(* Logix 5000 project; controller _GigaDiscovery vendor 1 type 14 code 244 rev 35.11; software revision 35.03; part 3 of 23 *)
(* tags used below, declared in another part *)
   Emergencies_Std_CL0 : DINT[8];
   Emergencies_Std_CL1 : DINT[8];
   Emergency_Captr : DINT[11];
   Fault_2_4 : Powerflex_DC_Fault;
   Fault_7 : Powerflex_DC_Fault;
   HMI_Drive_Fault_Descr : STRING[4];
   I_ADSL_Fault_Ch1 : BOOL;   // Gondola Communication Modem Fault CH1 -T27002C
   I_ADSL_Fault_Ch2 : BOOL;   // Gondola Communication Modem Fault CH2 -T27002C
   I_Compressor_Motor_Protection : BOOL;   // Compressor Motor Protection Feedback -F18002C
   I_Dryer_Motor_Protection : BOOL;   // Dryer Motor Protection Feedback -F18202C
   I_MCC_Temperature_OK : BOOL;   // MCC temeprature OK -S75003C
   I_Motor_1_2_Fan_Protection_Feedback : BOOL;   // Motor 1-2 Fan Protection Feedback -F10402C -F10406C
   I_Motor_1_Overvoltage_Control : BOOL;   // Motor 1 Overvoltage control - Relay OK -K10302G
   I_Motor_1_Thermal_Probe : BOOL;   // Motor 1 Thermal Probe -K10702H
   I_Motor_2_Overvoltage_Control : BOOL;   // Motor 2 Overvoltage control - Relay OK -K10307G
   I_Motor_2_Thermal_Probe : BOOL;   // Motor 2 Thermal Probe -K10704H
   I_Motor_3_4_Fan_Protection_Feedback : BOOL;   // Motor 3-4 Fan Protection Feedback -F12402C -F12406C
   I_Motor_3_Overvoltage_Control : BOOL;   // Motor 3 Overvoltage control - Relay OK -K12302G
   I_Motor_3_Thermal_Probe : BOOL;   // Motor 3 Thermal Probe -K12702H
   I_Motor_4_Overvoltage_Control : BOOL;   // Motor 4 Overvoltage control - Relay OK -K12307G
   I_Motor_4_Thermal_Probe : BOOL;   // Motor 4 Thermal Probe -K12704H
   I_Motor_5_6_Fan_Protection_Feedback : BOOL;   // Motor 5-6 Fan Protection Feedback -F14402C -F14406C
   I_Motor_5_Overvoltage_Control : BOOL;   // Motor 5 Overvoltage control - Relay OK -K14302G
   I_Motor_5_Thermal_Probe : BOOL;   // Motor 5 Thermal Probe -K14702H
   I_Motor_6_Overvoltage_Control : BOOL;   // Motor 6 Overvoltage control - Relay OK -K14307G
   I_Motor_6_Thermal_Probe : BOOL;   // Motor 6 Thermal Probe -K14704H
   I_Motor_7_Fan_Protection_Feedback : BOOL;   // Motor 7 Fan Protection Feedback -F16402C
   I_Motor_7_Thermal_Probe : BOOL;   // Motor 7 Thermal Probe -K16602H
   I_Pylon_Home_Ch1 : UDT_DCM;   // Home position Pylon Ch1 -B26002I
   I_Pylon_Home_Ch2 : UDT_DCM;   // Home position Pylon Ch2 -B26007I
   Jerk_Time : REAL;   // T1 Region 1
   PltaformClosed_CycleComplete : BOOL;   // Piattaforme chiuse e ciclo completato
   PltaformOpeneded_CycleComplete : BOOL;   // Rilevazione Piattaforme aperte con ciclo Completato
   Power_On_Delay : BOOL;
   Pylon_Axe : Axe;
   Real : REAL[32];
   Reset_Pulse : BOOL;
   RESTRAINTS_Rack_Sector_ON : BOOL;

        [6].I_Close_Position.ChannelA := 1, [6].I_Close_Position.ChannelB := 1, [6].I_Close_Position.InputStatus := 1, [6].I_Close_Position.SafetyFunction := 41, [6].I_Close_Position.DiscrepancyTime := 3000, [6].I_Close_Position.O1 := 1, [6].I_Close_Position.IS := 1, [6].I_Sector_Disable_Switch.Dual_Chanel_Monitor.ChannelB := 1, [6].I_Sector_Disable_Switch.Dual_Chanel_Monitor.InputStatus := 1, [6].I_Sector_Disable_Switch.Dual_Chanel_Monitor.SafetyFunction := 41, [6].I_Sector_Disable_Switch.Dual_Chanel_Monitor.InputType := 2, [6].I_Sector_Disable_Switch.Dual_Chanel_Monitor.DiscrepancyTime := 3000, [6].I_Sector_Disable_Switch.Dual_Chanel_Monitor.IS := 1, [6].I_Sector_Disable_Switch.Status := 1, [6].O_Unlock_Valve_Left.FeedBack_Type := 1, [6].O_Unlock_Valve_Left.Discrepancy_Time := 3000, [6].O_Unlock_Valve_Left.I_FeedBack_Data := 1, [6].O_Unlock_Valve_Left.I_FeedBack_Status := 1, [6].O_Unlock_Valve_Left.I_Output_Status := 1, [6].O_Unlock_Valve_Right.FeedBack_Type := 1, [6].O_Unlock_Valve_Right.Discrepancy_Time := 3000, [6].O_Unlock_Valve_Right.I_FeedBack_Data := 1, [6].O_Unlock_Valve_Right.I_FeedBack_Status := 1, [6].O_Unlock_Valve_Right.I_Output_Status := 1, [7].Sensors_ChA := 1, [7].Sensors_ChB := 1, [7].LapBar_Open_Close := 1, [7].Input_Status := 1, [7].Sensor_ChA_Open_Memory := 1, [7].Sensor_ChB_Open_Memory := 1, [7].I_LB_PressureSwitch_Valve_Right_Open := 1, [7].I_LB_PressureSwitch_Valve_Left_Open := 1, [7].All_Rack_Memory_Signal_ON := 1, [7].RESTRAINTS_Rack_Sector_ON := 1, [7].I_Close_Position.ChannelA := 1, [7].I_Close_Position.ChannelB := 1, [7].I_Close_Position.InputStatus := 1, [7].I_Close_Position.SafetyFunction := 41, [7].I_Close_Position.DiscrepancyTime := 3000, [7].I_Close_Position.O1 := 1, [7].I_Close_Position.IS := 1, [7].I_Sector_Disable_Switch.Dual_Chanel_Monitor.ChannelB := 1, [7].I_Sector_Disable_Switch.Dual_Chanel_Monitor.InputStatus := 1, [7].I_Sector_Disable_Switch.Dual_Chanel_Monitor.SafetyFunction := 41, [7].I_Sector_Disable_Switch.Dual_Chanel_Monitor.InputType := 2, [7].I_Sector_Disable_Switch.Dual_Chanel_Monitor.DiscrepancyTime := 3000, [7].I_Sector_Disable_Switch.Dual_Chanel_Monitor.IS := 1, [7].I_Sector_Disable_Switch.Status := 1, [7].O_Unlock_Valve_Left.FeedBack_Type := 1, [7].O_Unlock_Valve_Left.Discrepancy_Time := 3000, [7].O_Unlock_Valve_Left.I_FeedBack_Data := 1, [7].O_Unlock_Valve_Left.I_FeedBack_Status := 1, [7].O_Unlock_Valve_Left.I_Output_Status := 1, [7].O_Unlock_Valve_Right.FeedBack_Type := 1, [7].O_Unlock_Valve_Right.Discrepancy_Time := 3000, [7].O_Unlock_Valve_Right.I_FeedBack_Data := 1, [7].O_Unlock_Valve_Right.I_FeedBack_Status := 1, [7].O_Unlock_Valve_Right.I_Output_Status := 1, [8].Sensors_ChA := 1, [8].Sensors_ChB := 1,
        [8].LapBar_Open_Close := 1, [8].Input_Status := 1, [8].Sensor_ChA_Open_Memory := 1, [8].Sensor_ChB_Open_Memory := 1, [8].I_LB_PressureSwitch_Valve_Right_Open := 1, [8].I_LB_PressureSwitch_Valve_Left_Open := 1, [8].All_Rack_Memory_Signal_ON := 1, [8].RESTRAINTS_Rack_Sector_ON := 1, [8].I_Close_Position.ChannelA := 1, [8].I_Close_Position.ChannelB := 1, [8].I_Close_Position.InputStatus := 1, [8].I_Close_Position.SafetyFunction := 41, [8].I_Close_Position.DiscrepancyTime := 3000, [8].I_Close_Position.O1 := 1, [8].I_Close_Position.IS := 1, [8].I_Sector_Disable_Switch.Dual_Chanel_Monitor.ChannelB := 1, [8].I_Sector_Disable_Switch.Dual_Chanel_Monitor.InputStatus := 1, [8].I_Sector_Disable_Switch.Dual_Chanel_Monitor.SafetyFunction := 41, [8].I_Sector_Disable_Switch.Dual_Chanel_Monitor.InputType := 2, [8].I_Sector_Disable_Switch.Dual_Chanel_Monitor.DiscrepancyTime := 3000, [8].I_Sector_Disable_Switch.Dual_Chanel_Monitor.IS := 1, [8].I_Sector_Disable_Switch.Status := 1, [8].O_Unlock_Valve_Left.FeedBack_Type := 1, [8].O_Unlock_Valve_Left.Discrepancy_Time := 3000, [8].O_Unlock_Valve_Left.I_FeedBack_Data := 1, [8].O_Unlock_Valve_Left.I_FeedBack_Status := 1, [8].O_Unlock_Valve_Left.I_Output_Status := 1, [8].O_Unlock_Valve_Right.FeedBack_Type := 1, [8].O_Unlock_Valve_Right.Discrepancy_Time := 3000, [8].O_Unlock_Valve_Right.I_FeedBack_Data := 1, [8].O_Unlock_Valve_Right.I_FeedBack_Status := 1, [8].O_Unlock_Valve_Right.I_Output_Status := 1);
        [1].I_Sector_Disable_Switch   // -DOOR-S27802F SECTOR A ENABLE
        [2].I_Sector_Disable_Switch   // -DOOR-S27806F SECTOR B ENABLE
        [3].I_Sector_Disable_Switch   // -DOOR-S27902F SECTOR C ENABLE
        [4].I_Sector_Disable_Switch   // -DOOR-S27906F SECTOR D ENABLE
        [5].I_Sector_Disable_Switch   // -DOOR-S28002F SECTOR E ENABLE
        [6].I_Sector_Disable_Switch   // -DOOR-S28006F SECTOR F ENABLE
        [7].I_Sector_Disable_Switch   // -DOOR-S28102F SECTOR G ENABLE
        [8].I_Sector_Disable_Switch   // -DOOR-S28106F SECTOR H ENABLE
        [3]   // Lapbars Sector C Seats 11 to 15
        [1].I_LB_PressureSwitch_Valve_Left_Open   // -S50602J
        [1].I_LB_PressureSwitch_Valve_Right_Open   // -S50606J
        [2].I_LB_PressureSwitch_Valve_Left_Open   // -S52602J
        [2].I_LB_PressureSwitch_Valve_Right_Open   // -S52606J
        [3].I_LB_PressureSwitch_Valve_Left_Open   // -S54602J
        [3].I_LB_PressureSwitch_Valve_Right_Open   // -S54606J
        [4].I_LB_PressureSwitch_Valve_Left_Open   // -S56602J
        [4].I_LB_PressureSwitch_Valve_Right_Open   // -S56606J
        [5].I_LB_PressureSwitch_Valve_Left_Open   // -S58602J
        [5].I_LB_PressureSwitch_Valve_Right_Open   // -S58606J
        [6].I_LB_PressureSwitch_Valve_Left_Open   // -S60602J
        [6].I_LB_PressureSwitch_Valve_Right_Open   // -S60606J
        [7].I_LB_PressureSwitch_Valve_Left_Open   // -S62602J
        [7].I_LB_PressureSwitch_Valve_Right_Open   // -S62606J
        [8].I_LB_PressureSwitch_Valve_Left_Open   // -S64602J
        [8].I_LB_PressureSwitch_Valve_Right_Open   // -S64606J
        [4]   // Lapbars Sector D Seats 16 to 20
        [6]   // Lapbars Sector F Seats 26 to 30
        [2]   // Lapbars Sector B Seats 6 to 10
        [5]   // Lapbars Sector E Seats 21 to25
        [7]   // Lapbars Sector G Seats 31 to 35
        [8]   // Lapbars Sector H Seats 36 to 40
        [1]   // Lapbars Sector A Seats 1 to 5
   RESTRAINTS_Sector_Enable_OFF : BOOL := 1;   // ALL RESTRAINTS rack commands OFF
   RESTRAINTS_Sector_Enable_ON : BOOL;   // ALL RESTRAINTS Sector Enable ON
   RESTRAINTS_Unlock_Valve_Pressure : BOOL := 1;
   Revolution_time_1 : DINT := 15480;
   Revolution_time_2 : DINT := 15520;
   RPM_Max_Motor_Speed_Pylon : DINT := 1710;
   SCP_K : STD_SCP := (Input := 13.991667, Input_Max := 14.0, Input_Min := 12.0, Output := -3.0083332, Scaled_Max := -3.0, Scaled_Min := -5.0);
   SCuve_K_Stop : S_Curve_Calc := (Jerk_Time := 1.0, Accel_Time := 3.0, Jerk_Rate := 25.0, Accel_Rate := 25.0);
   Second_Oscillation_Done : BOOL;   // Second Oscillation End
   SEL_T3_R011 : SELECT;
   SEL_T3_R0112 : SELECT;
   Speed_at_Minute : REAL := 928.8;
   Speed_at_Second : REAL := 15.48;
   Speed_Treshold : REAL := 10.0;
   Start_Autom_Cycle : Sequencer := (Step_Timer[0].PRE := 5000, Step_Timer[0].ACC := 5000, Step_Timer[0].EN := 1, Step_Timer[0].DN := 1, Step_Timer[1].PRE := 500, Step_Timer[2].PRE := 6000, Step_Timer[3].PRE := 20000, Step_Timer[3].ACC := 20000, Step_Timer[3].DN := 1, Step_Timer[4].PRE := 500, Step_Timer[4].ACC := 500, Step_Timer[4].EN := 1, Step_Timer[4].DN := 1, Step_Timer[5].PRE := 85000, Step_Timer[7].PRE := 1000, Step_Timer[8].PRE := 1000, Step_Timer[9].PRE := 500, Time_Limit[3].PRE := 40000, Time_Limit[8].PRE := 80000, Step_00 := 1);
        .Step_01   // Imposto velocità e verso di marcia rotazione gondola RST arms homming
        .Step_03   // Fase di Stop del pilone e rallentamento gondla
        .Step_09   // Stop disalimento il teleruttore di marcia
        .Step_04   // Imposto la velocità vicino allo Zero
        .Step_02   // Avvio Oscillazione pilone
        .Step_08   // Stop disabilito il drive della Gondola
        .Step_20   // Fast Stop
        .Step_07   // Stop
   Start_Permissive : Permissive := (BitsConditions := -269484034);
   Start_Permissive2 : Permissive := (BitsConditions := -8);
   Start_Platform_AutoCycle_Pylon : BOOL;
   Start_Stop_Cycle : Sequencer := (Step_Timer[0].PRE := 1000, Step_Timer[1].PRE := 500, Step_Timer[2].PRE := 500, Step_Timer[3].PRE := 1000, Step_Timer[4].PRE := 500, Step_Timer[8].PRE := 200, Time_Limit[1].PRE := 2000, Time_Limit[2].PRE := 2000, Time_Limit[3].PRE := 2000, Time_Limit[4].PRE := 2000, Time_Limit[5].PRE := 5000, Time_Limit[6].PRE := 2000, Time_Limit[7].PRE := 2000, Time_Limit[8].PRE := 10000, Time_Limit[9].PRE := 50000, Time_Limit[10].PRE := 7000, Step_00 := 1);
        .Step_28   // 28 Disalimento i teleruttori di potenza dei drive
        .Step_04   // Accendo Teleruttori per il Campo dei Motori 5 (Gondola)
        .Step_02   // Accendo Teleruttori per lo Start e per il Campo dei Drive (pylon)
        .Step_01   // I start opening the platforms
        .Step_15   // Disabilito i Drive
        .Step_06   // Abilito la Potenza
        .Step_09   // Disabilito i Drive
        .Step_07   // Abilito i convertitori
        .Step_12   // Tolgo lo start e metto lo stop ai drive
        .Step_08   // Comando lo Start ai convertitori
        .Step_31   // Cycle Ended
        .Step_10   // Avvio le oscillazioni della giostra
   Start_TOF : TIMER := (PRE := 5000, ACC := 5000);
   Stats_Times : DINT[30] := ([1] := 231);
        [10]   // encoder difference?
        [1]   // Time Run Started
   Stop_K_to_Zero : BOOL;
   Stop_Request : BOOL;
   Target_Angle : REAL := 120.0;
   Test : DCI_STOP_TEST;
   TimeInStation_Count_Daily : COUNTER := (PRE := 500, ACC := 6);
   TimeInStation_Count_Hourly : COUNTER := (PRE := 100, ACC := 2);
   TimeInStation_Timer : TIMER := (PRE := 600000);   // 10 min 600 sec
   Timer_Overspeed_reset_1 : BOOL;   // senor 1 Revolution time reset
   Timer_Overspeed_reset_2 : BOOL;   // senor 2
   Timers : TIMER[32] := ([0].PRE := 300, [0].ACC := 300, [1].PRE := 1000, [2].PRE := 60000, [3].PRE := 10000, [4].PRE := 10000, [5].PRE := 2000, [6].PRE := 10000, [7].PRE := 1000, [8].PRE := 200, [9].PRE := 200, [10].PRE := 10000, [11].PRE := 1000, [12].PRE := 2500, [13].PRE := 1000, [14].PRE := 10000, [15].PRE := 10000, [16].PRE := 2000, [16].ACC := 2000, [17].PRE := 2000, [18].PRE := 2000, [19].PRE := 1000, [20].PRE := 100, [21].PRE := 100, [22].PRE := 100, [23].PRE := 1000, [24].PRE := 500, [24].ACC := 130, [24].EN := 1, [24].TT := 1, [25].PRE := 500, [26].PRE := 125, [26].ACC := 18, [26].EN := 1, [26].TT := 1, [27].PRE := 125, [28].PRE := 2000, [29].PRE := 2000, [29].ACC := 2001, [29].EN := 1, [29].DN := 1, [30].PRE := 2000, [31].PRE := 10000, [31].ACC := 10001, [31].EN := 1, [31].DN := 1);
   To_Sfty : Std_to_Sfty := (Seat_Auxiliary_Ch_Memory := 1, I_Fan_Feedback_NO := 1, RFID_Reset := 1, No_Std_Emergencies_CL0 := 1, No_Std_Emergencies_CL1 := 1, Pylon_min_speed := 1, Gondola_min_Speed := 1, Fbk_MainCotnactor_M1_M3 := 1, Fbk_MainContactor_M2_M4 := 1, I_Gondola_Field_Contactor_Fdbk := 1, I_Gondola_Fuse_Power_Supply := 1, Motors_Temperature_Ok := 1, Low_speed_thold_emergency_brake := 1, UPS_RCC.I_Alarm := 1, UPS_RCC.O_Control := 1, UPS_MCC.I_Alarm := 1, UPS_MCC.O_Control := 1, Main_valve_Time := 10, HMI_Page := 400, Date_Time.Year := 2025, Date_Time.Month := 12, Date_Time.Day := 1, Date_Time.Hour := 19, Date_Time.Minute := 40, Date_Time.Second := 53, Date_Time.Milli_sec := 807892);
        .I_Fan_Feedback_NO   // Fan Feedback NO Pag.94
        .I_Fan_Feedback_NC   // Fan Feedback NC Pag.94
        .Fbk_PylonBrake_Contactor   // Pylon Brake Command Feedback -Q10801E
        .I_Magnalock_4_Closed   // Magnalock Gate 4 - Status Lock -A25307I
        .I_Magnalock_3_Closed   // Magnalock Gate 3 - Status Lock -A25301I
        .I_Magnalock_2_Closed   // Magnalock Gate 2 - Status Lock -A25207I
        .I_Magnalock_1_Closed   // Magnalock Gate 1 - Status Lock -A25201I
        .I_OCC2_Alarms_Reset_Pb   // OCC02 Reset FAult S6310E (Pag.86A)
   ToBe_Define_Sfty : DINT[10] := ([0] := -2147481679, [1] := -1);
        [0].10   // Verificare se va bene la logica per l'attivazione dle campo a riposo
   TobeDefine : DINT := 25;
   Torque_Cmd_from_Cycle : REAL;
   Torque_Filter : REAL := 7.0;
   Torque_To_Zero_Stewp_04 : BOOL;
   TorqueNeg_Angle_Control : REAL := -20.0;
   TorquePos_Angle_Control : REAL := 77.39982;
   Valve_Proof_Test_Cycle : Sequencer := (Step_Timer[0].PRE := 1000, Step_Timer[1].PRE := 2000, Step_Timer[2].PRE := 2000, Step_00 := 1);
        .Step_05   // Activate Close Platform Valve
        .Step_31   // Valve Proof Test Successful
        .Step_04   // Activate Open Platform Valve
        .Step_00   // Sequencer Stopped
        .Step_01   // Activate Main and close Valves
        .Step_02   // Verify that there's no pressure in the Open/Close Line
        .Step_03   // Turn OFF Main Valve
   Valve_Proof_Test_Ok : BOOL;
   Valve_Test_AOI : Sequencer_AOI;
   Valves_Pressure_Discrepancy : DINT := 3000;
   Warning : DINT[10];
        [0].1   // Gondola Communication Modem Fault CH1 -T27002C
        [0].2   // Gondola Communication Modem Fault CH2 -T27002C
        [0].0   // Gate Selector Switch Turned during cycle
        [0].5   // Dryer Motor Protection Feedback -F18202C
   Work_Auto_Cycle : Auto_Cycle := (Pylon_Angle := 120, Cycle_Time_min := 2, Cycle_Time_sec := 25, Gondola_Speed[0] := 20, Gondola_Speed[1] := 70, Gondola_Speed[2] := -75, Gondola_Speed[3] := 50, Gondola_Time[1] := 60, Gondola_Time[2] := 50, Gondola_Time[3] := 20);
   Work_Auto_Cycle_Ptr : DINT := 1;
END_VAR

PROGRAM Alarms   (* main routine Main *)
VAR
   Alarm_Timers : TIMER[64] := ([0].PRE := 300000, [1].PRE := 1000, [1].ACC := 1000, [2].PRE := 60000, [3].PRE := 60000, [4].PRE := 1000, [5].PRE := 1000, [6].PRE := 1000, [7].PRE := 1000, [8].PRE := 1000, [9].PRE := 300000, [10].PRE := 2000, [11].PRE := 10000, [12].PRE := 10000, [13].PRE := 5000, [14].PRE := 4000, [15].PRE := 4500, [16].PRE := 60000, [16].ACC := 60004, [16].EN := 1, [16].DN := 1, [17].PRE := 20000, [18].PRE := 1000, [18].ACC := 1000, [19].PRE := 1000, [19].ACC := 1000, [20].PRE := 500, [21].PRE := 4000, [22].PRE := 250, [22].EN := 1, [23].PRE := 250, [24].PRE := 500, [24].ACC := 502, [25].PRE := 1500, [25].ACC := 1500, [26].PRE := 300, [27].PRE := 1000, [27].ACC := 1000, [27].EN := 1, [27].DN := 1, [28].PRE := 3000, [28].ACC := 3001, [28].EN := 1, [28].DN := 1, [29].PRE := 1000, [30].PRE := 1000, [31].PRE := 1000, [32].PRE := 60000, [32].ACC := 60004, [32].EN := 1, [32].DN := 1, [33].PRE := 1800000);
        [25]   // Larghezza impulso di reset Convertitori
   Fault_1_3 : Powerflex_DC_Fault := (Fault_Code := 75);
   Fault_5_6 : Powerflex_DC_Fault := (Fault_Code := 75);
   Os : DINT;
        .0   // USED
        .1   // USED
        .2   // USED
        .3   // USED
        .4   // USED
        .5   // USED
END_VAR

ROUTINE _00_Alarm_Manage   (* ladder *)
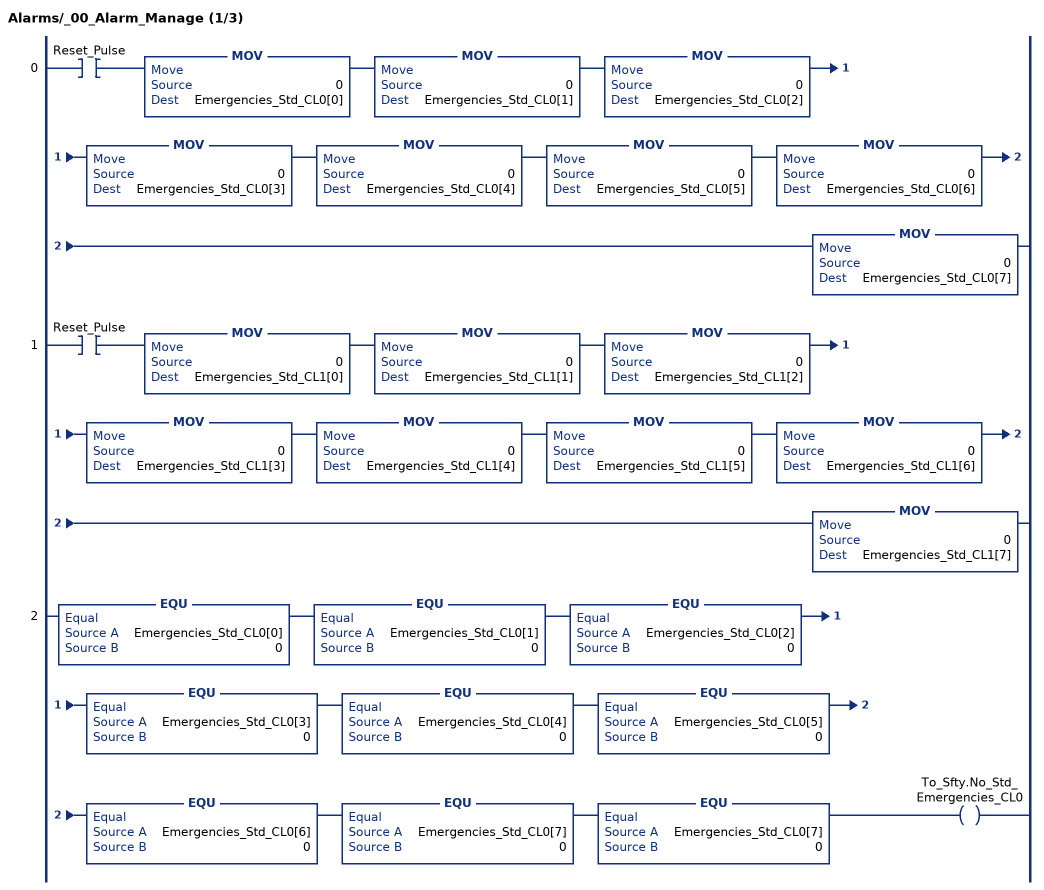
   0: XIC(Reset_Pulse)MOV(0,Emergencies_Std_CL0[0])MOV(0,Emergencies_Std_CL0[1])MOV(0,Emergencies_Std_CL0[2])MOV(0,Emergencies_Std_CL0[3])MOV(0,Emergencies_Std_CL0[4])MOV(0,Emergencies_Std_CL0[5])MOV(0,Emergencies_Std_CL0[6])MOV(0,Emergencies_Std_CL0[7]);
   1: XIC(Reset_Pulse)MOV(0,Emergencies_Std_CL1[0])MOV(0,Emergencies_Std_CL1[1])MOV(0,Emergencies_Std_CL1[2])MOV(0,Emergencies_Std_CL1[3])MOV(0,Emergencies_Std_CL1[4])MOV(0,Emergencies_Std_CL1[5])MOV(0,Emergencies_Std_CL1[6])MOV(0,Emergencies_Std_CL1[7]);
   2: EQU(Emergencies_Std_CL0[0],0)EQU(Emergencies_Std_CL0[1],0)EQU(Emergencies_Std_CL0[2],0)EQU(Emergencies_Std_CL0[3],0)EQU(Emergencies_Std_CL0[4],0)EQU(Emergencies_Std_CL0[5],0)EQU(Emergencies_Std_CL0[6],0)EQU(Emergencies_Std_CL0[7],0)EQU(Emergencies_Std_CL0[7],0)OTE(To_Sfty.No_Std_Emergencies_CL0);
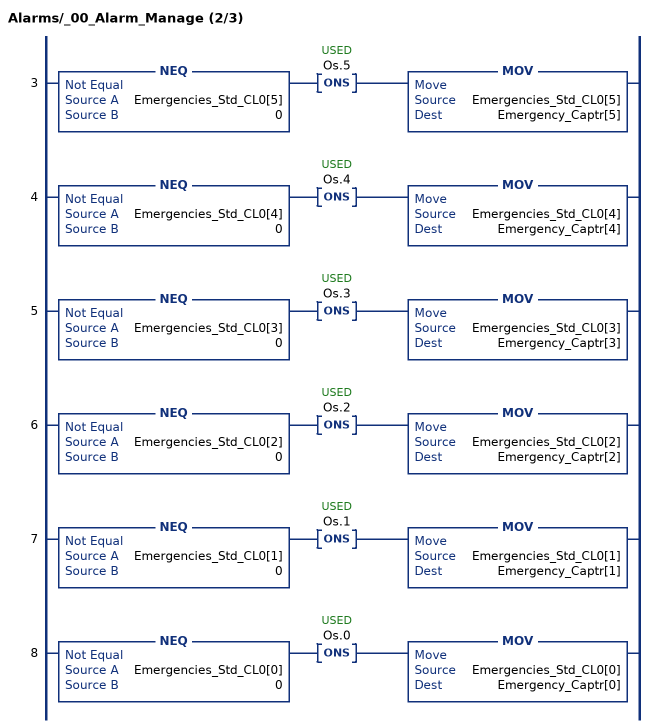
   3: NEQ(Emergencies_Std_CL0[5],0)ONS(Os.5)MOV(Emergencies_Std_CL0[5],Emergency_Captr[5]);
   4: NEQ(Emergencies_Std_CL0[4],0)ONS(Os.4)MOV(Emergencies_Std_CL0[4],Emergency_Captr[4]);
   5: NEQ(Emergencies_Std_CL0[3],0)ONS(Os.3)MOV(Emergencies_Std_CL0[3],Emergency_Captr[3]);
   6: NEQ(Emergencies_Std_CL0[2],0)ONS(Os.2)MOV(Emergencies_Std_CL0[2],Emergency_Captr[2]);
   7: NEQ(Emergencies_Std_CL0[1],0)ONS(Os.1)MOV(Emergencies_Std_CL0[1],Emergency_Captr[1]);
   8: NEQ(Emergencies_Std_CL0[0],0)ONS(Os.0)MOV(Emergencies_Std_CL0[0],Emergency_Captr[0]);
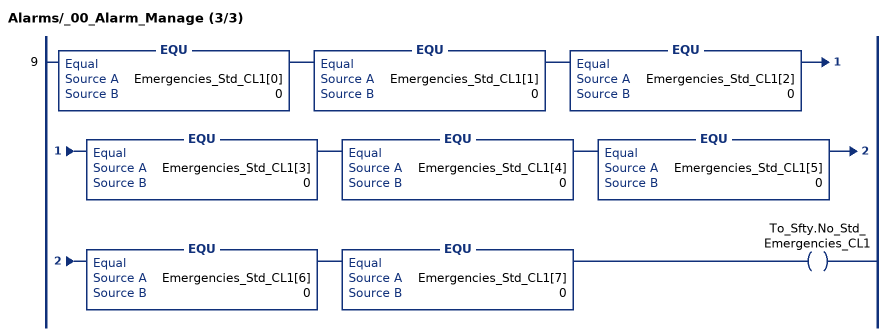
   9: EQU(Emergencies_Std_CL1[0],0)EQU(Emergencies_Std_CL1[1],0)EQU(Emergencies_Std_CL1[2],0)EQU(Emergencies_Std_CL1[3],0)EQU(Emergencies_Std_CL1[4],0)EQU(Emergencies_Std_CL1[5],0)EQU(Emergencies_Std_CL1[6],0)EQU(Emergencies_Std_CL1[7],0)OTE(To_Sfty.No_Std_Emergencies_CL1);
END_ROUTINE

ROUTINE _01_MCC   (* ladder *)
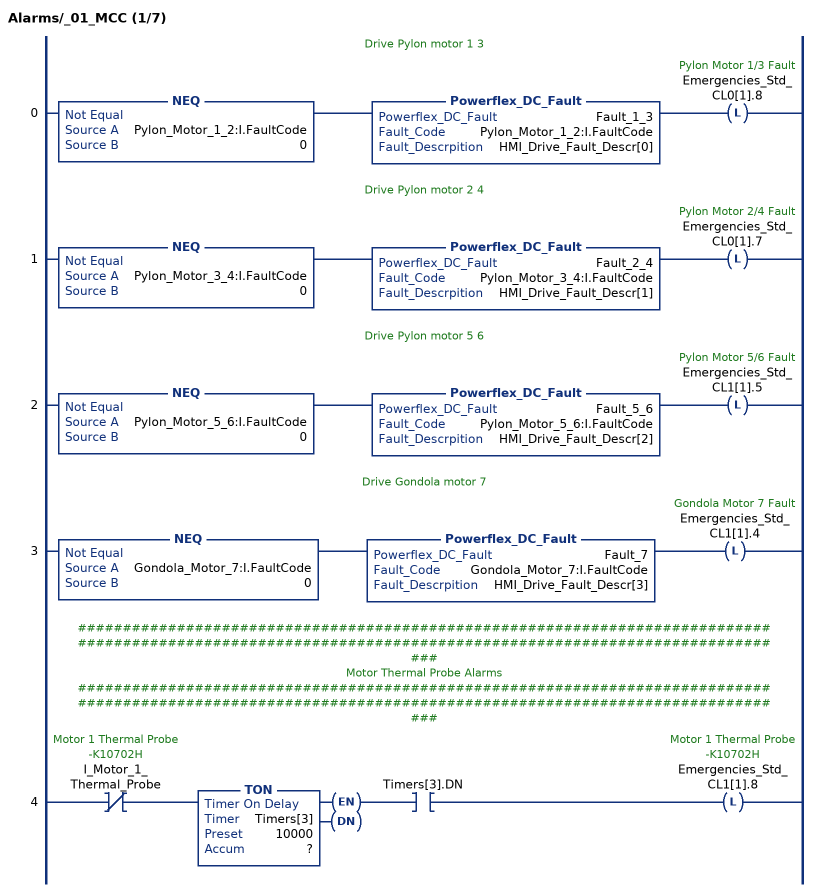
   // Drive Pylon motor 1 3
   0: NEQ(Pylon_Motor_1_2:I.FaultCode,0)Powerflex_DC_Fault(Fault_1_3,Pylon_Motor_1_2:I.FaultCode,HMI_Drive_Fault_Descr[0])OTL(Emergencies_Std_CL0[1].8);
   // Drive Pylon motor 2 4
   1: NEQ(Pylon_Motor_3_4:I.FaultCode,0)Powerflex_DC_Fault(Fault_2_4,Pylon_Motor_3_4:I.FaultCode,HMI_Drive_Fault_Descr[1])OTL(Emergencies_Std_CL0[1].7);
   // Drive Pylon motor 5 6
   2: NEQ(Pylon_Motor_5_6:I.FaultCode,0)Powerflex_DC_Fault(Fault_5_6,Pylon_Motor_5_6:I.FaultCode,HMI_Drive_Fault_Descr[2])OTL(Emergencies_Std_CL1[1].5);
   // Drive Gondola motor 7
   3: NEQ(Gondola_Motor_7:I.FaultCode,0)Powerflex_DC_Fault(Fault_7,Gondola_Motor_7:I.FaultCode,HMI_Drive_Fault_Descr[3])OTL(Emergencies_Std_CL1[1].4);
   // #############################################################################################################################################################
   // Motor Thermal Probe Alarms
   // #############################################################################################################################################################
   4: XIO(I_Motor_1_Thermal_Probe)TON(Timers[3],?,?)XIC(Timers[3].DN)OTL(Emergencies_Std_CL1[1].8);
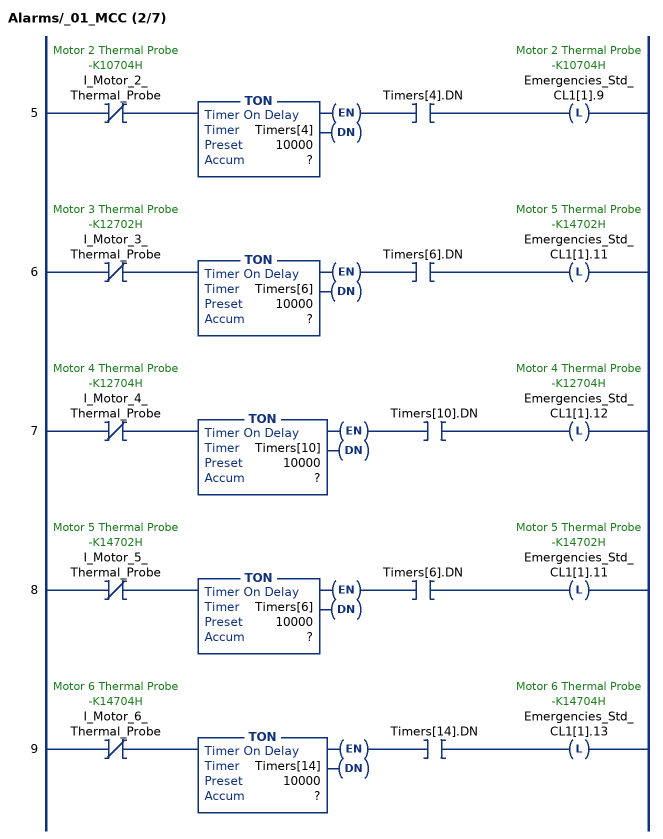
   5: XIO(I_Motor_2_Thermal_Probe)TON(Timers[4],?,?)XIC(Timers[4].DN)OTL(Emergencies_Std_CL1[1].9);
   6: XIO(I_Motor_3_Thermal_Probe)TON(Timers[6],?,?)XIC(Timers[6].DN)OTL(Emergencies_Std_CL1[1].11);
   7: XIO(I_Motor_4_Thermal_Probe)TON(Timers[10],?,?)XIC(Timers[10].DN)OTL(Emergencies_Std_CL1[1].12);
   8: XIO(I_Motor_5_Thermal_Probe)TON(Timers[6],?,?)XIC(Timers[6].DN)OTL(Emergencies_Std_CL1[1].11);
   9: XIO(I_Motor_6_Thermal_Probe)TON(Timers[14],?,?)XIC(Timers[14].DN)OTL(Emergencies_Std_CL1[1].13);
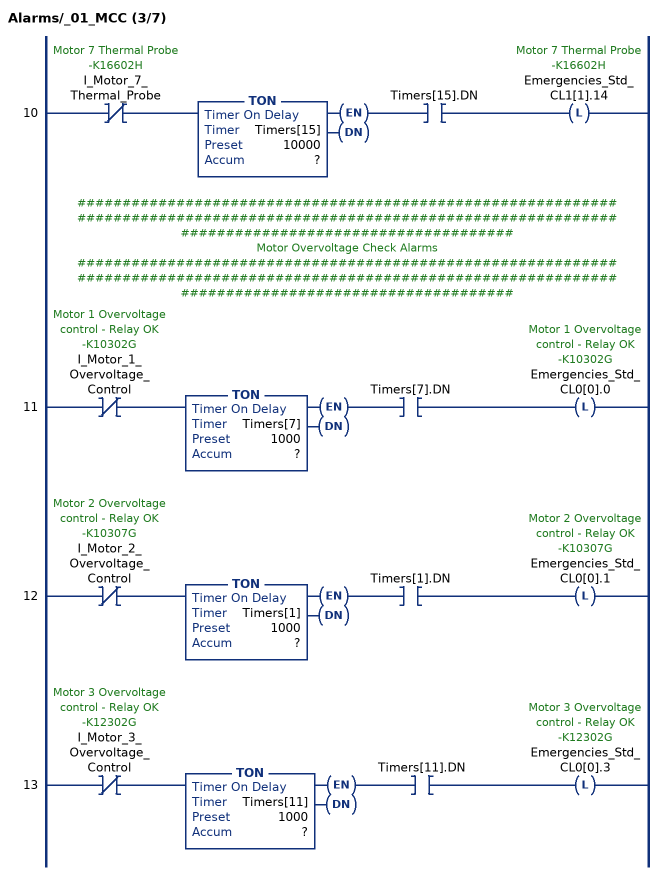
   10: XIO(I_Motor_7_Thermal_Probe)TON(Timers[15],?,?)XIC(Timers[15].DN)OTL(Emergencies_Std_CL1[1].14);
   // #############################################################################################################################################################
   // Motor Overvoltage Check Alarms
   // #############################################################################################################################################################
   11: XIO(I_Motor_1_Overvoltage_Control)TON(Timers[7],?,?)XIC(Timers[7].DN)OTL(Emergencies_Std_CL0[0].0);
   12: XIO(I_Motor_2_Overvoltage_Control)TON(Timers[1],?,?)XIC(Timers[1].DN)OTL(Emergencies_Std_CL0[0].1);
   13: XIO(I_Motor_3_Overvoltage_Control)TON(Timers[11],?,?)XIC(Timers[11].DN)OTL(Emergencies_Std_CL0[0].3);
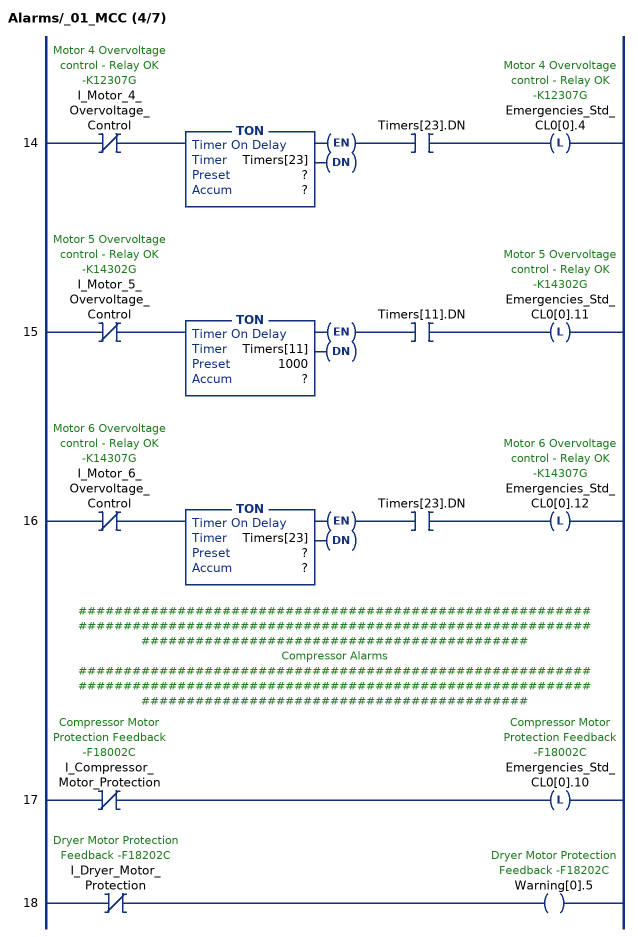
   14: XIO(I_Motor_4_Overvoltage_Control)TON(Timers[23],?,?)XIC(Timers[23].DN)OTL(Emergencies_Std_CL0[0].4);
   15: XIO(I_Motor_5_Overvoltage_Control)TON(Timers[11],?,?)XIC(Timers[11].DN)OTL(Emergencies_Std_CL0[0].11);
   16: XIO(I_Motor_6_Overvoltage_Control)TON(Timers[23],?,?)XIC(Timers[23].DN)OTL(Emergencies_Std_CL0[0].12);
   // #############################################################################################################################################################
   // Compressor Alarms
   // #############################################################################################################################################################
   17: XIO(I_Compressor_Motor_Protection)OTL(Emergencies_Std_CL0[0].10);
   18: XIO(I_Dryer_Motor_Protection)OTE(Warning[0].5);
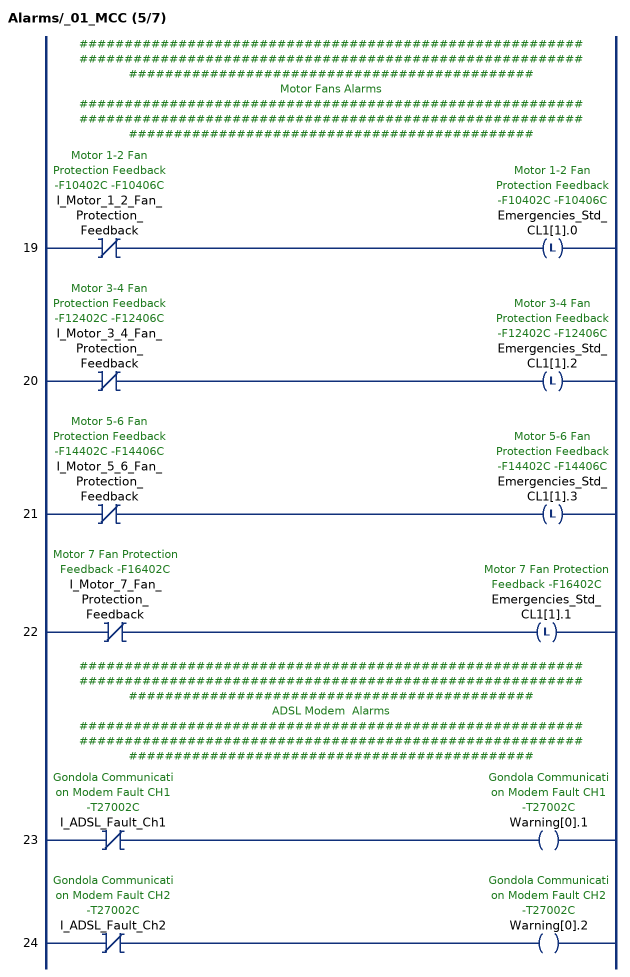
   // #############################################################################################################################################################
   // Motor Fans Alarms
   // #############################################################################################################################################################
   19: XIO(I_Motor_1_2_Fan_Protection_Feedback)OTL(Emergencies_Std_CL1[1].0);
   20: XIO(I_Motor_3_4_Fan_Protection_Feedback)OTL(Emergencies_Std_CL1[1].2);
   21: XIO(I_Motor_5_6_Fan_Protection_Feedback)OTL(Emergencies_Std_CL1[1].3);
   22: XIO(I_Motor_7_Fan_Protection_Feedback)OTL(Emergencies_Std_CL1[1].1);
   // #############################################################################################################################################################
   // ADSL Modem  Alarms
   // #############################################################################################################################################################
   23: XIO(I_ADSL_Fault_Ch1)OTE(Warning[0].1);
   24: XIO(I_ADSL_Fault_Ch2)OTE(Warning[0].2);
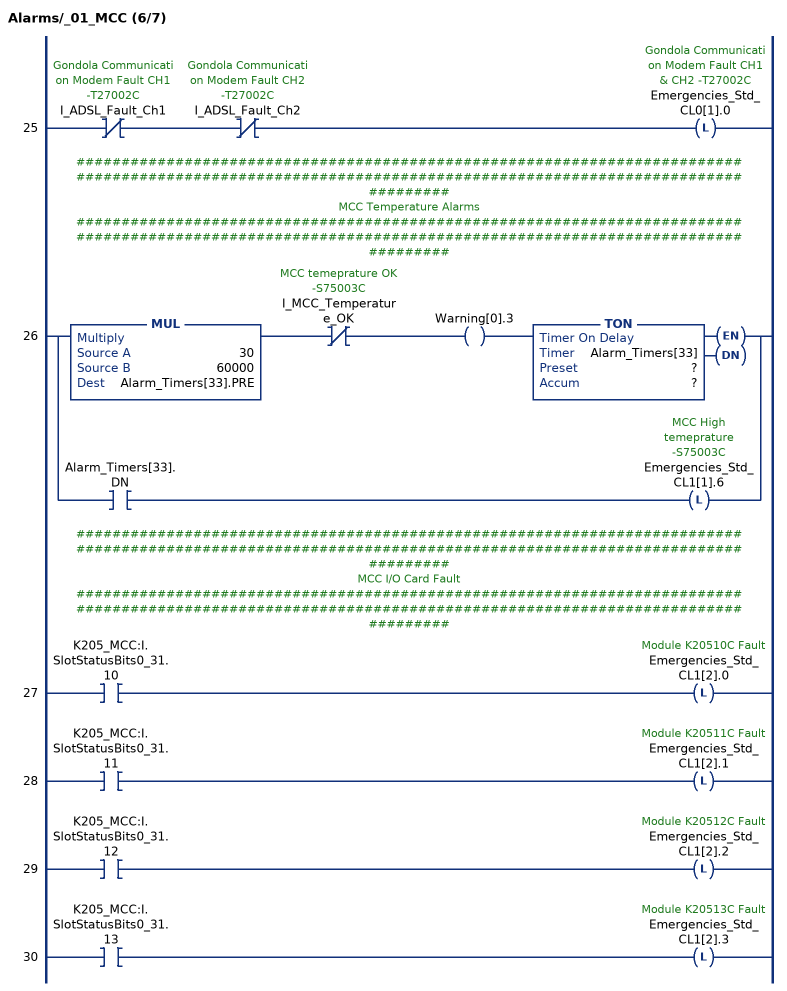
   25: XIO(I_ADSL_Fault_Ch1)XIO(I_ADSL_Fault_Ch2)OTL(Emergencies_Std_CL0[1].0);
   // #############################################################################################################################################################
   // MCC Temperature Alarms
   // #############################################################################################################################################################
   26: [MUL(30,60000,Alarm_Timers[33].PRE) XIO(I_MCC_Temperature_OK) OTE(Warning[0].3) TON(Alarm_Timers[33],?,?) ,XIC(Alarm_Timers[33].DN) OTL(Emergencies_Std_CL1[1].6) ];
   // #############################################################################################################################################################
   // MCC I/O Card Fault
   // #############################################################################################################################################################
   27: XIC(K205_MCC:I.SlotStatusBits0_31.10)OTL(Emergencies_Std_CL1[2].0);
   28: XIC(K205_MCC:I.SlotStatusBits0_31.11)OTL(Emergencies_Std_CL1[2].1);
   29: XIC(K205_MCC:I.SlotStatusBits0_31.12)OTL(Emergencies_Std_CL1[2].2);
   30: XIC(K205_MCC:I.SlotStatusBits0_31.13)OTL(Emergencies_Std_CL1[2].3);
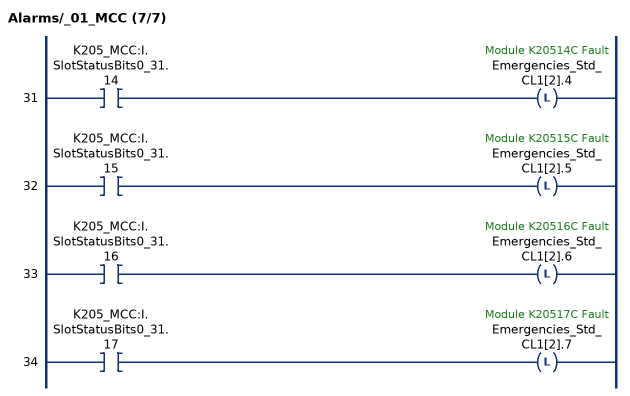
   31: XIC(K205_MCC:I.SlotStatusBits0_31.14)OTL(Emergencies_Std_CL1[2].4);
   32: XIC(K205_MCC:I.SlotStatusBits0_31.15)OTL(Emergencies_Std_CL1[2].5);
   33: XIC(K205_MCC:I.SlotStatusBits0_31.16)OTL(Emergencies_Std_CL1[2].6);
   34: XIC(K205_MCC:I.SlotStatusBits0_31.17)OTL(Emergencies_Std_CL1[2].7);
END_ROUTINE

ROUTINE _04_Pylon   (* ladder *)